REGION Network 12: IW422 - Tank Group Pressure (PT-424) - Tank Group
   RUNG wire#powerrail
      { S7_Templates := "[SrcType := Int, DestType := Real]" } Normalize(min := "20_TANKS_IP_DATA".RIO_07.FIRST_TANK.TANKS_PRESS_CNFG.RAW_MIN, value := "RIO7 Tank Pressure", max := "20_TANKS_IP_DATA".RIO_07.FIRST_TANK.TANKS_PRESS_CNFG.RAW_MAX, out => "20_TANKS_IP_DATA".RIO_07.FIRST_TANK.TANKS_PRESS_CNFG.NORM)
      { S7_Templates := "[SrcType := Real, DestType := Real]" } Scale(min := "20_TANKS_IP_DATA".RIO_07.FIRST_TANK.TANKS_PRESS_CNFG.ENG_MIN, value := "20_TANKS_IP_DATA".RIO_07.FIRST_TANK.TANKS_PRESS_CNFG.NORM, max := "20_TANKS_IP_DATA".RIO_07.FIRST_TANK.TANKS_PRESS_CNFG.ENG_MAX, out => "20_TANKS_IP_DATA".RIO_07.FIRST_TANK.TANKS_PRESS)
   END_RUNG
   // the same network as SCL:
   "20_TANKS_IP_DATA".RIO_07.FIRST_TANK.TANKS_PRESS_CNFG.NORM := NORM_X(MIN := "20_TANKS_IP_DATA".RIO_07.FIRST_TANK.TANKS_PRESS_CNFG.RAW_MIN, VALUE := "RIO7 Tank Pressure", MAX := "20_TANKS_IP_DATA".RIO_07.FIRST_TANK.TANKS_PRESS_CNFG.RAW_MAX);
   "20_TANKS_IP_DATA".RIO_07.FIRST_TANK.TANKS_PRESS := SCALE_X(MIN := "20_TANKS_IP_DATA".RIO_07.FIRST_TANK.TANKS_PRESS_CNFG.ENG_MIN, VALUE := "20_TANKS_IP_DATA".RIO_07.FIRST_TANK.TANKS_PRESS_CNFG.NORM, MAX := "20_TANKS_IP_DATA".RIO_07.FIRST_TANK.TANKS_PRESS_CNFG.ENG_MAX);
END_REGION
END_FUNCTION

FUNCTION "40_RIO_Output_Processing" : Void   // FC40, LAD
TITLE = RIO Output Processing
{ S7_Optimized_Access := 'TRUE' }
AUTHOR : JRS
VERSION : 0.1
// To call output processing blocks in logical order
BEGIN

REGION Network 1: RIO Digital Output Processing - Rack 1
   // To process code outputs prior to physical connection
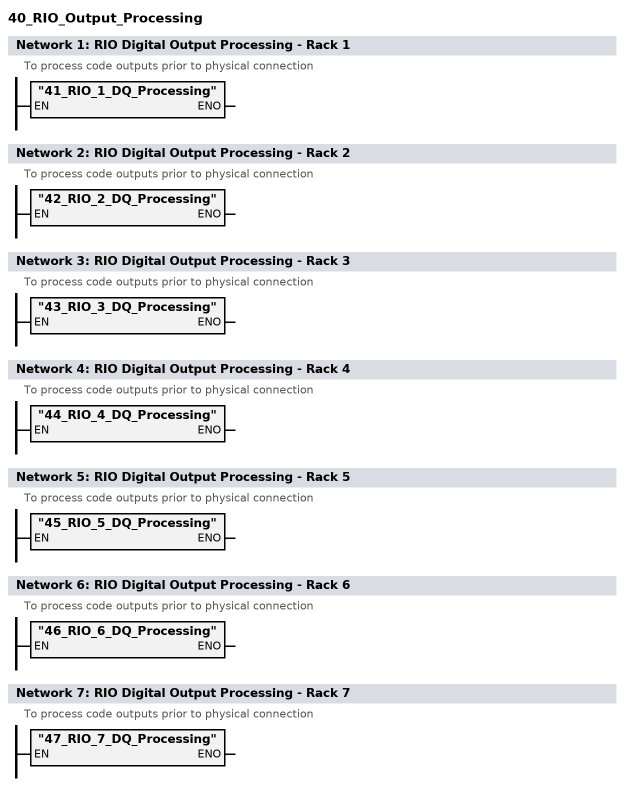
   RUNG wire#powerrail
      "41_RIO_1_DQ_Processing"()
   END_RUNG
   // the same network as SCL:
   "41_RIO_1_DQ_Processing"();
END_REGION

REGION Network 2: RIO Digital Output Processing - Rack 2
   // To process code outputs prior to physical connection
   RUNG wire#powerrail
      "42_RIO_2_DQ_Processing"()
   END_RUNG
   // the same network as SCL:
   "42_RIO_2_DQ_Processing"();
END_REGION

REGION Network 3: RIO Digital Output Processing - Rack 3
   // To process code outputs prior to physical connection
   RUNG wire#powerrail
      "43_RIO_3_DQ_Processing"()
   END_RUNG
   // the same network as SCL:
   "43_RIO_3_DQ_Processing"();
END_REGION

REGION Network 4: RIO Digital Output Processing - Rack 4
   // To process code outputs prior to physical connection
   RUNG wire#powerrail
      "44_RIO_4_DQ_Processing"()
   END_RUNG
   // the same network as SCL:
   "44_RIO_4_DQ_Processing"();
END_REGION

REGION Network 5: RIO Digital Output Processing - Rack 5
   // To process code outputs prior to physical connection
   RUNG wire#powerrail
      "45_RIO_5_DQ_Processing"()
   END_RUNG
   // the same network as SCL:
   "45_RIO_5_DQ_Processing"();
END_REGION

REGION Network 6: RIO Digital Output Processing - Rack 6
   // To process code outputs prior to physical connection
   RUNG wire#powerrail
      "46_RIO_6_DQ_Processing"()
   END_RUNG
   // the same network as SCL:
   "46_RIO_6_DQ_Processing"();
END_REGION

REGION Network 7: RIO Digital Output Processing - Rack 7
   // To process code outputs prior to physical connection
   RUNG wire#powerrail
      "47_RIO_7_DQ_Processing"()
   END_RUNG
   // the same network as SCL:
   "47_RIO_7_DQ_Processing"();
END_REGION
END_FUNCTION

FUNCTION "41_RIO_1_DQ_Processing" : Void   // FC41, LAD
TITLE = RIO Rack Digital Output Processing (Tanks APT, 1P & 1S)
{ S7_Optimized_Access := 'TRUE' }
AUTHOR : JRS
VERSION : 0.1
// To process code outputs prior to physical connection
BEGIN

REGION Network 1: Q0.0 - Tank Vent Valve Control (CV-441-A) - FPT
   // True = CLOSE, False = OPEN
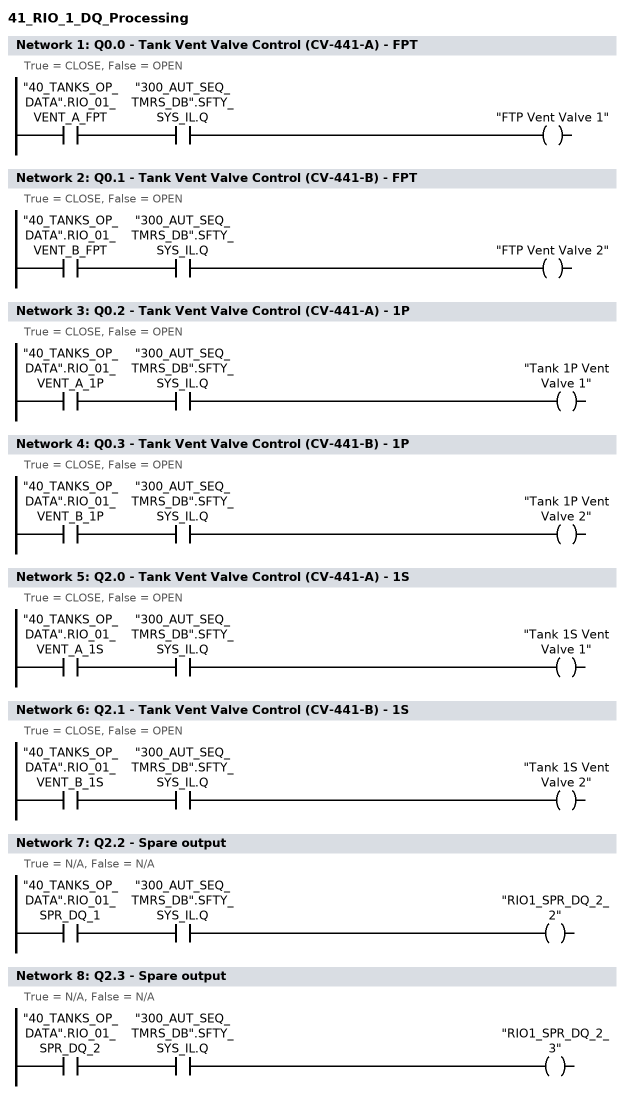
   RUNG wire#powerrail
      Contact( "40_TANKS_OP_DATA".RIO_01_VENT_A_FPT )
      Contact( "300_AUT_SEQ_TMRS_DB".SFTY_SYS_IL.Q )
      Coil( "FTP Vent Valve 1" )
   END_RUNG
   // the same network as SCL:
   "FTP Vent Valve 1" := "40_TANKS_OP_DATA".RIO_01_VENT_A_FPT AND "300_AUT_SEQ_TMRS_DB".SFTY_SYS_IL.Q;
END_REGION

REGION Network 2: Q0.1 - Tank Vent Valve Control (CV-441-B) - FPT
   // True = CLOSE, False = OPEN
   RUNG wire#powerrail
      Contact( "40_TANKS_OP_DATA".RIO_01_VENT_B_FPT )
      Contact( "300_AUT_SEQ_TMRS_DB".SFTY_SYS_IL.Q )
      Coil( "FTP Vent Valve 2" )
   END_RUNG
   // the same network as SCL:
   "FTP Vent Valve 2" := "40_TANKS_OP_DATA".RIO_01_VENT_B_FPT AND "300_AUT_SEQ_TMRS_DB".SFTY_SYS_IL.Q;
END_REGION

REGION Network 3: Q0.2 - Tank Vent Valve Control (CV-441-A) - 1P
   // True = CLOSE, False = OPEN
   RUNG wire#powerrail
      Contact( "40_TANKS_OP_DATA".RIO_01_VENT_A_1P )
      Contact( "300_AUT_SEQ_TMRS_DB".SFTY_SYS_IL.Q )
      Coil( "Tank 1P Vent Valve 1" )
   END_RUNG
   // the same network as SCL:
   "Tank 1P Vent Valve 1" := "40_TANKS_OP_DATA".RIO_01_VENT_A_1P AND "300_AUT_SEQ_TMRS_DB".SFTY_SYS_IL.Q;
END_REGION

REGION Network 4: Q0.3 - Tank Vent Valve Control (CV-441-B) - 1P
   // True = CLOSE, False = OPEN
   RUNG wire#powerrail
      Contact( "40_TANKS_OP_DATA".RIO_01_VENT_B_1P )
      Contact( "300_AUT_SEQ_TMRS_DB".SFTY_SYS_IL.Q )
      Coil( "Tank 1P Vent Valve 2" )
   END_RUNG
   // the same network as SCL:
   "Tank 1P Vent Valve 2" := "40_TANKS_OP_DATA".RIO_01_VENT_B_1P AND "300_AUT_SEQ_TMRS_DB".SFTY_SYS_IL.Q;
END_REGION

REGION Network 5: Q2.0 - Tank Vent Valve Control (CV-441-A) - 1S
   // True = CLOSE, False = OPEN
   RUNG wire#powerrail
      Contact( "40_TANKS_OP_DATA".RIO_01_VENT_A_1S )
      Contact( "300_AUT_SEQ_TMRS_DB".SFTY_SYS_IL.Q )
      Coil( "Tank 1S Vent Valve 1" )
   END_RUNG
   // the same network as SCL:
   "Tank 1S Vent Valve 1" := "40_TANKS_OP_DATA".RIO_01_VENT_A_1S AND "300_AUT_SEQ_TMRS_DB".SFTY_SYS_IL.Q;
END_REGION

REGION Network 6: Q2.1 - Tank Vent Valve Control (CV-441-B) - 1S
   // True = CLOSE, False = OPEN
   RUNG wire#powerrail
      Contact( "40_TANKS_OP_DATA".RIO_01_VENT_B_1S )
      Contact( "300_AUT_SEQ_TMRS_DB".SFTY_SYS_IL.Q )
      Coil( "Tank 1S Vent Valve 2" )
   END_RUNG
   // the same network as SCL:
   "Tank 1S Vent Valve 2" := "40_TANKS_OP_DATA".RIO_01_VENT_B_1S AND "300_AUT_SEQ_TMRS_DB".SFTY_SYS_IL.Q;
END_REGION

REGION Network 7: Q2.2 - Spare output
   // True = N/A, False = N/A
   RUNG wire#powerrail
      Contact( "40_TANKS_OP_DATA".RIO_01_SPR_DQ_1 )
      Contact( "300_AUT_SEQ_TMRS_DB".SFTY_SYS_IL.Q )
      Coil( "RIO1_SPR_DQ_2_2" )
   END_RUNG
   // the same network as SCL:
   "RIO1_SPR_DQ_2_2" := "40_TANKS_OP_DATA".RIO_01_SPR_DQ_1 AND "300_AUT_SEQ_TMRS_DB".SFTY_SYS_IL.Q;
END_REGION

REGION Network 8: Q2.3 - Spare output
   // True = N/A, False = N/A
   RUNG wire#powerrail
      Contact( "40_TANKS_OP_DATA".RIO_01_SPR_DQ_2 )
      Contact( "300_AUT_SEQ_TMRS_DB".SFTY_SYS_IL.Q )
      Coil( "RIO1_SPR_DQ_2_3" )
   END_RUNG
   // the same network as SCL:
   "RIO1_SPR_DQ_2_3" := "40_TANKS_OP_DATA".RIO_01_SPR_DQ_2 AND "300_AUT_SEQ_TMRS_DB".SFTY_SYS_IL.Q;
END_REGION
END_FUNCTION

FUNCTION "42_RIO_2_DQ_Processing" : Void   // FC42, LAD
TITLE = RIO Rack Digital Output Processing (Tanks 2P & 2S)
{ S7_Optimized_Access := 'TRUE' }
AUTHOR : JRS
VERSION : 0.1
// To process code outputs prior to physical connection
BEGIN

REGION Network 1: Q6.0 - Tank Vent Valve Control (CV-441-A) - 2P
   // True = CLOSE, False = OPEN
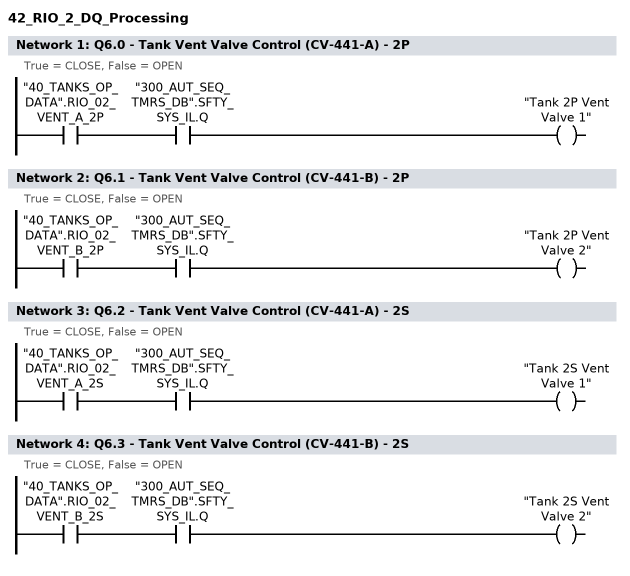
   RUNG wire#powerrail
      Contact( "40_TANKS_OP_DATA".RIO_02_VENT_A_2P )
      Contact( "300_AUT_SEQ_TMRS_DB".SFTY_SYS_IL.Q )
      Coil( "Tank 2P Vent Valve 1" )
   END_RUNG
   // the same network as SCL:
   "Tank 2P Vent Valve 1" := "40_TANKS_OP_DATA".RIO_02_VENT_A_2P AND "300_AUT_SEQ_TMRS_DB".SFTY_SYS_IL.Q;
END_REGION

REGION Network 2: Q6.1 - Tank Vent Valve Control (CV-441-B) - 2P
   // True = CLOSE, False = OPEN
   RUNG wire#powerrail
      Contact( "40_TANKS_OP_DATA".RIO_02_VENT_B_2P )
      Contact( "300_AUT_SEQ_TMRS_DB".SFTY_SYS_IL.Q )
      Coil( "Tank 2P Vent Valve 2" )
   END_RUNG
   // the same network as SCL:
   "Tank 2P Vent Valve 2" := "40_TANKS_OP_DATA".RIO_02_VENT_B_2P AND "300_AUT_SEQ_TMRS_DB".SFTY_SYS_IL.Q;
END_REGION

REGION Network 3: Q6.2 - Tank Vent Valve Control (CV-441-A) - 2S
   // True = CLOSE, False = OPEN
   RUNG wire#powerrail
      Contact( "40_TANKS_OP_DATA".RIO_02_VENT_A_2S )
      Contact( "300_AUT_SEQ_TMRS_DB".SFTY_SYS_IL.Q )
      Coil( "Tank 2S Vent Valve 1" )
   END_RUNG
   // the same network as SCL:
   "Tank 2S Vent Valve 1" := "40_TANKS_OP_DATA".RIO_02_VENT_A_2S AND "300_AUT_SEQ_TMRS_DB".SFTY_SYS_IL.Q;
END_REGION

REGION Network 4: Q6.3 - Tank Vent Valve Control (CV-441-B) - 2S
   // True = CLOSE, False = OPEN
   RUNG wire#powerrail
      Contact( "40_TANKS_OP_DATA".RIO_02_VENT_B_2S )
      Contact( "300_AUT_SEQ_TMRS_DB".SFTY_SYS_IL.Q )
      Coil( "Tank 2S Vent Valve 2" )
   END_RUNG
   // the same network as SCL:
   "Tank 2S Vent Valve 2" := "40_TANKS_OP_DATA".RIO_02_VENT_B_2S AND "300_AUT_SEQ_TMRS_DB".SFTY_SYS_IL.Q;
END_REGION
END_FUNCTION

FUNCTION "43_RIO_3_DQ_Processing" : Void   // FC43, LAD
TITLE = RIO Rack Digital Output Processing (Tanks 3P & 3S)
{ S7_Optimized_Access := 'TRUE' }
AUTHOR : JRS
VERSION : 0.1
// To process code outputs prior to physical connection
BEGIN

REGION Network 1: Q10.0 - Tank Vent Valve Control (CV-441-A) - 3P
   // True = CLOSE, False = OPEN
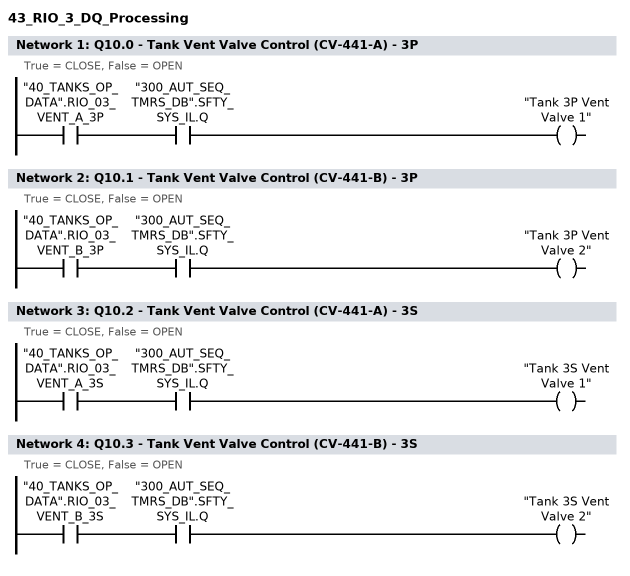
   RUNG wire#powerrail
      Contact( "40_TANKS_OP_DATA".RIO_03_VENT_A_3P )
      Contact( "300_AUT_SEQ_TMRS_DB".SFTY_SYS_IL.Q )
      Coil( "Tank 3P Vent Valve 1" )
   END_RUNG
   // the same network as SCL:
   "Tank 3P Vent Valve 1" := "40_TANKS_OP_DATA".RIO_03_VENT_A_3P AND "300_AUT_SEQ_TMRS_DB".SFTY_SYS_IL.Q;
END_REGION

REGION Network 2: Q10.1 - Tank Vent Valve Control (CV-441-B) - 3P
   // True = CLOSE, False = OPEN
   RUNG wire#powerrail
      Contact( "40_TANKS_OP_DATA".RIO_03_VENT_B_3P )
      Contact( "300_AUT_SEQ_TMRS_DB".SFTY_SYS_IL.Q )
      Coil( "Tank 3P Vent Valve 2" )
   END_RUNG
   // the same network as SCL:
   "Tank 3P Vent Valve 2" := "40_TANKS_OP_DATA".RIO_03_VENT_B_3P AND "300_AUT_SEQ_TMRS_DB".SFTY_SYS_IL.Q;
END_REGION

REGION Network 3: Q10.2 - Tank Vent Valve Control (CV-441-A) - 3S
   // True = CLOSE, False = OPEN
   RUNG wire#powerrail
      Contact( "40_TANKS_OP_DATA".RIO_03_VENT_A_3S )
      Contact( "300_AUT_SEQ_TMRS_DB".SFTY_SYS_IL.Q )
      Coil( "Tank 3S Vent Valve 1" )
   END_RUNG
   // the same network as SCL:
   "Tank 3S Vent Valve 1" := "40_TANKS_OP_DATA".RIO_03_VENT_A_3S AND "300_AUT_SEQ_TMRS_DB".SFTY_SYS_IL.Q;
END_REGION

REGION Network 4: Q10.3 - Tank Vent Valve Control (CV-441-B) - 3S
   // True = CLOSE, False = OPEN
   RUNG wire#powerrail
      Contact( "40_TANKS_OP_DATA".RIO_03_VENT_B_3S )
      Contact( "300_AUT_SEQ_TMRS_DB".SFTY_SYS_IL.Q )
      Coil( "Tank 3S Vent Valve 2" )
   END_RUNG
   // the same network as SCL:
   "Tank 3S Vent Valve 2" := "40_TANKS_OP_DATA".RIO_03_VENT_B_3S AND "300_AUT_SEQ_TMRS_DB".SFTY_SYS_IL.Q;
END_REGION
END_FUNCTION

FUNCTION "44_RIO_4_DQ_Processing" : Void   // FC44, LAD
TITLE = RIO Rack Digital Output Processing (Tanks 4P & 4S)
{ S7_Optimized_Access := 'TRUE' }
AUTHOR : JRS
VERSION : 0.1
// To process code outputs prior to physical connection
BEGIN

REGION Network 1: Q14.0 - Tank Vent Valve Control (CV-441-A) - 4P
   // True = CLOSE, False = OPEN
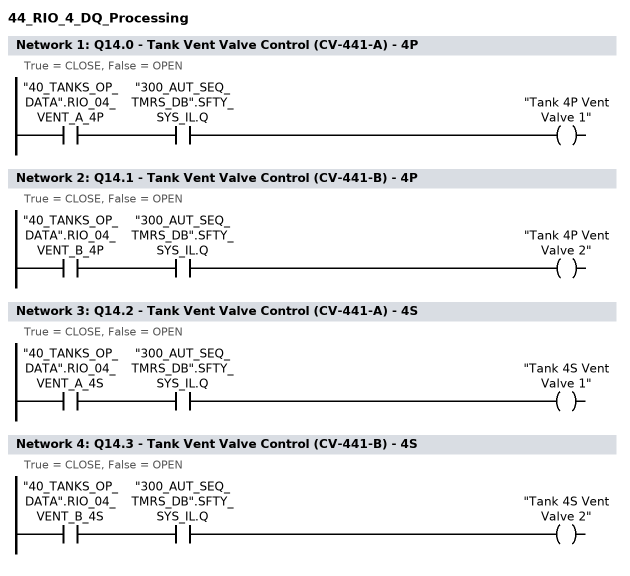
   RUNG wire#powerrail
      Contact( "40_TANKS_OP_DATA".RIO_04_VENT_A_4P )
      Contact( "300_AUT_SEQ_TMRS_DB".SFTY_SYS_IL.Q )
      Coil( "Tank 4P Vent Valve 1" )
   END_RUNG
   // the same network as SCL:
   "Tank 4P Vent Valve 1" := "40_TANKS_OP_DATA".RIO_04_VENT_A_4P AND "300_AUT_SEQ_TMRS_DB".SFTY_SYS_IL.Q;
END_REGION

REGION Network 2: Q14.1 - Tank Vent Valve Control (CV-441-B) - 4P
   // True = CLOSE, False = OPEN
   RUNG wire#powerrail
      Contact( "40_TANKS_OP_DATA".RIO_04_VENT_B_4P )
      Contact( "300_AUT_SEQ_TMRS_DB".SFTY_SYS_IL.Q )
      Coil( "Tank 4P Vent Valve 2" )
   END_RUNG
   // the same network as SCL:
   "Tank 4P Vent Valve 2" := "40_TANKS_OP_DATA".RIO_04_VENT_B_4P AND "300_AUT_SEQ_TMRS_DB".SFTY_SYS_IL.Q;
END_REGION

REGION Network 3: Q14.2 - Tank Vent Valve Control (CV-441-A) - 4S
   // True = CLOSE, False = OPEN
   RUNG wire#powerrail
      Contact( "40_TANKS_OP_DATA".RIO_04_VENT_A_4S )
      Contact( "300_AUT_SEQ_TMRS_DB".SFTY_SYS_IL.Q )
      Coil( "Tank 4S Vent Valve 1" )
   END_RUNG
   // the same network as SCL:
   "Tank 4S Vent Valve 1" := "40_TANKS_OP_DATA".RIO_04_VENT_A_4S AND "300_AUT_SEQ_TMRS_DB".SFTY_SYS_IL.Q;
END_REGION

REGION Network 4: Q14.3 - Tank Vent Valve Control (CV-441-B) - 4S
   // True = CLOSE, False = OPEN
   RUNG wire#powerrail
      Contact( "40_TANKS_OP_DATA".RIO_04_VENT_B_4S )
      Contact( "300_AUT_SEQ_TMRS_DB".SFTY_SYS_IL.Q )
      Coil( "Tank 4S Vent Valve 2" )
   END_RUNG
   // the same network as SCL:
   "Tank 4S Vent Valve 2" := "40_TANKS_OP_DATA".RIO_04_VENT_B_4S AND "300_AUT_SEQ_TMRS_DB".SFTY_SYS_IL.Q;
END_REGION
END_FUNCTION

FUNCTION "45_RIO_5_DQ_Processing" : Void   // FC45, LAD
TITLE = RIO Rack Digital Output Processing (Tanks 5P & 5S)
{ S7_Optimized_Access := 'TRUE' }
AUTHOR : JRS
VERSION : 0.1
// To process code outputs prior to physical connection
BEGIN

REGION Network 1: Q18.0 - Tank Vent Valve Control (CV-441-A) - 5P
   // True = CLOSE, False = OPEN
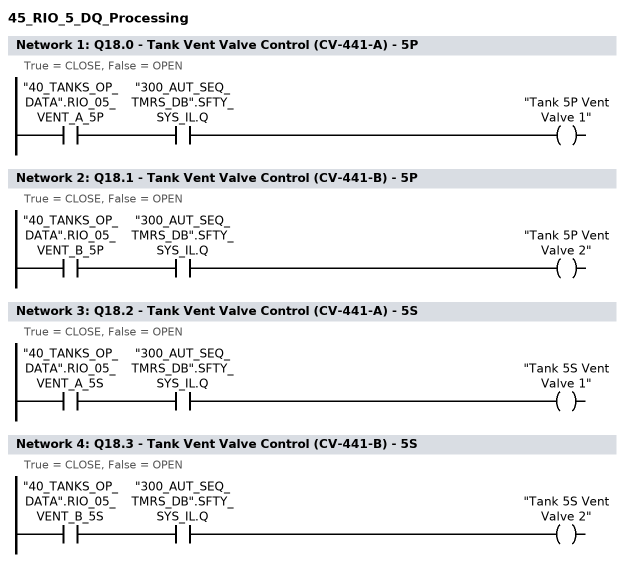
   RUNG wire#powerrail
      Contact( "40_TANKS_OP_DATA".RIO_05_VENT_A_5P )
      Contact( "300_AUT_SEQ_TMRS_DB".SFTY_SYS_IL.Q )
      Coil( "Tank 5P Vent Valve 1" )
   END_RUNG
   // the same network as SCL:
   "Tank 5P Vent Valve 1" := "40_TANKS_OP_DATA".RIO_05_VENT_A_5P AND "300_AUT_SEQ_TMRS_DB".SFTY_SYS_IL.Q;
END_REGION

REGION Network 2: Q18.1 - Tank Vent Valve Control (CV-441-B) - 5P
   // True = CLOSE, False = OPEN
   RUNG wire#powerrail
      Contact( "40_TANKS_OP_DATA".RIO_05_VENT_B_5P )
      Contact( "300_AUT_SEQ_TMRS_DB".SFTY_SYS_IL.Q )
      Coil( "Tank 5P Vent Valve 2" )
   END_RUNG
   // the same network as SCL:
   "Tank 5P Vent Valve 2" := "40_TANKS_OP_DATA".RIO_05_VENT_B_5P AND "300_AUT_SEQ_TMRS_DB".SFTY_SYS_IL.Q;
END_REGION

REGION Network 3: Q18.2 - Tank Vent Valve Control (CV-441-A) - 5S
   // True = CLOSE, False = OPEN
   RUNG wire#powerrail
      Contact( "40_TANKS_OP_DATA".RIO_05_VENT_A_5S )
      Contact( "300_AUT_SEQ_TMRS_DB".SFTY_SYS_IL.Q )
      Coil( "Tank 5S Vent Valve 1" )
   END_RUNG
   // the same network as SCL:
   "Tank 5S Vent Valve 1" := "40_TANKS_OP_DATA".RIO_05_VENT_A_5S AND "300_AUT_SEQ_TMRS_DB".SFTY_SYS_IL.Q;
END_REGION

REGION Network 4: Q18.3 - Tank Vent Valve Control (CV-441-B) - 5S
   // True = CLOSE, False = OPEN
   RUNG wire#powerrail
      Contact( "40_TANKS_OP_DATA".RIO_05_VENT_B_5S )
      Contact( "300_AUT_SEQ_TMRS_DB".SFTY_SYS_IL.Q )
      Coil( "Tank 5S Vent Valve 2" )
   END_RUNG
   // the same network as SCL:
   "Tank 5S Vent Valve 2" := "40_TANKS_OP_DATA".RIO_05_VENT_B_5S AND "300_AUT_SEQ_TMRS_DB".SFTY_SYS_IL.Q;
END_REGION
END_FUNCTION

FUNCTION "46_RIO_6_DQ_Processing" : Void   // FC46, LAD
TITLE = RIO Rack Digital Output Processing (Tanks 6P & 6S)
{ S7_Optimized_Access := 'TRUE' }
AUTHOR : JRS
VERSION : 0.1
// To process code outputs prior to physical connection
BEGIN

REGION Network 1: Q20.0 - Tank Vent Valve Control (CV-441-A) - 6P
   // True = CLOSE, False = OPEN
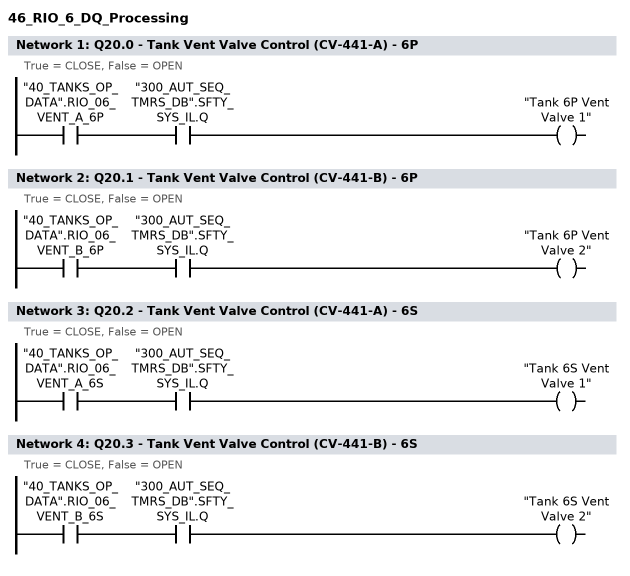
   RUNG wire#powerrail
      Contact( "40_TANKS_OP_DATA".RIO_06_VENT_A_6P )
      Contact( "300_AUT_SEQ_TMRS_DB".SFTY_SYS_IL.Q )
      Coil( "Tank 6P Vent Valve 1" )
   END_RUNG
   // the same network as SCL:
   "Tank 6P Vent Valve 1" := "40_TANKS_OP_DATA".RIO_06_VENT_A_6P AND "300_AUT_SEQ_TMRS_DB".SFTY_SYS_IL.Q;
END_REGION

REGION Network 2: Q20.1 - Tank Vent Valve Control (CV-441-B) - 6P
   // True = CLOSE, False = OPEN
   RUNG wire#powerrail
      Contact( "40_TANKS_OP_DATA".RIO_06_VENT_B_6P )
      Contact( "300_AUT_SEQ_TMRS_DB".SFTY_SYS_IL.Q )
      Coil( "Tank 6P Vent Valve 2" )
   END_RUNG
   // the same network as SCL:
   "Tank 6P Vent Valve 2" := "40_TANKS_OP_DATA".RIO_06_VENT_B_6P AND "300_AUT_SEQ_TMRS_DB".SFTY_SYS_IL.Q;
END_REGION

REGION Network 3: Q20.2 - Tank Vent Valve Control (CV-441-A) - 6S
   // True = CLOSE, False = OPEN
   RUNG wire#powerrail
      Contact( "40_TANKS_OP_DATA".RIO_06_VENT_A_6S )
      Contact( "300_AUT_SEQ_TMRS_DB".SFTY_SYS_IL.Q )
      Coil( "Tank 6S Vent Valve 1" )
   END_RUNG
   // the same network as SCL:
   "Tank 6S Vent Valve 1" := "40_TANKS_OP_DATA".RIO_06_VENT_A_6S AND "300_AUT_SEQ_TMRS_DB".SFTY_SYS_IL.Q;
END_REGION

REGION Network 4: Q20.3 - Tank Vent Valve Control (CV-441-B) - 6S
   // True = CLOSE, False = OPEN
   RUNG wire#powerrail
      Contact( "40_TANKS_OP_DATA".RIO_06_VENT_B_6S )
      Contact( "300_AUT_SEQ_TMRS_DB".SFTY_SYS_IL.Q )
      Coil( "Tank 6S Vent Valve 2" )
   END_RUNG
   // the same network as SCL:
   "Tank 6S Vent Valve 2" := "40_TANKS_OP_DATA".RIO_06_VENT_B_6S AND "300_AUT_SEQ_TMRS_DB".SFTY_SYS_IL.Q;
END_REGION
END_FUNCTION

FUNCTION "47_RIO_7_DQ_Processing" : Void   // FC47, LAD
TITLE = RIO Rack Digital Output Processing (Tank APT)
{ S7_Optimized_Access := 'TRUE' }
AUTHOR : JRS
VERSION : 0.1
// To process code outputs prior to physical connection
BEGIN

REGION Network 1: Q26.0 - Tank Vent Valve Control (CV-441-A) - APT
   // True = CLOSE, False = OPEN
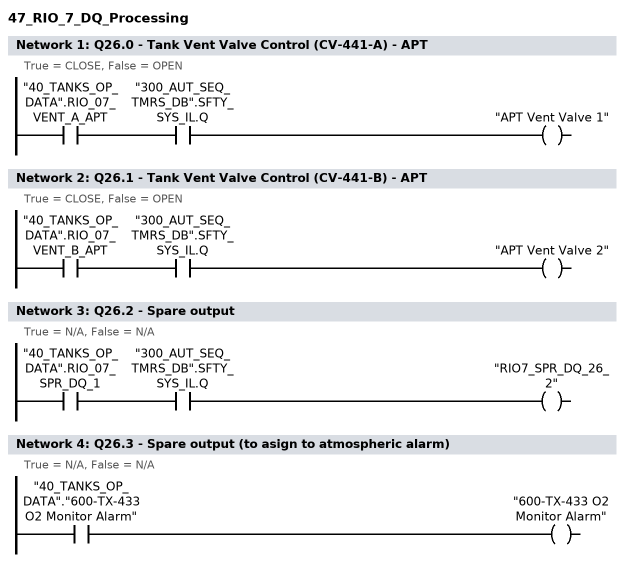
   RUNG wire#powerrail
      Contact( "40_TANKS_OP_DATA".RIO_07_VENT_A_APT )
      Contact( "300_AUT_SEQ_TMRS_DB".SFTY_SYS_IL.Q )
      Coil( "APT Vent Valve 1" )
   END_RUNG
   // the same network as SCL:
   "APT Vent Valve 1" := "40_TANKS_OP_DATA".RIO_07_VENT_A_APT AND "300_AUT_SEQ_TMRS_DB".SFTY_SYS_IL.Q;
END_REGION

REGION Network 2: Q26.1 - Tank Vent Valve Control (CV-441-B) - APT
   // True = CLOSE, False = OPEN
   RUNG wire#powerrail
      Contact( "40_TANKS_OP_DATA".RIO_07_VENT_B_APT )
      Contact( "300_AUT_SEQ_TMRS_DB".SFTY_SYS_IL.Q )
      Coil( "APT Vent Valve 2" )
   END_RUNG
   // the same network as SCL:
   "APT Vent Valve 2" := "40_TANKS_OP_DATA".RIO_07_VENT_B_APT AND "300_AUT_SEQ_TMRS_DB".SFTY_SYS_IL.Q;
END_REGION

REGION Network 3: Q26.2 - Spare output
   // True = N/A, False = N/A
   RUNG wire#powerrail
      Contact( "40_TANKS_OP_DATA".RIO_07_SPR_DQ_1 )
      Contact( "300_AUT_SEQ_TMRS_DB".SFTY_SYS_IL.Q )
      Coil( "RIO7_SPR_DQ_26_2" )
   END_RUNG
   // the same network as SCL:
   "RIO7_SPR_DQ_26_2" := "40_TANKS_OP_DATA".RIO_07_SPR_DQ_1 AND "300_AUT_SEQ_TMRS_DB".SFTY_SYS_IL.Q;
END_REGION

REGION Network 4: Q26.3 - Spare output (to asign to atmospheric alarm)
   // True = N/A, False = N/A
   RUNG wire#powerrail
      Contact( "40_TANKS_OP_DATA"."600-TX-433  O2 Monitor Alarm" )
      Coil( "600-TX-433 O2 Monitor Alarm" )
   END_RUNG
   // the same network as SCL:
   "600-TX-433 O2 Monitor Alarm" := "40_TANKS_OP_DATA"."600-TX-433  O2 Monitor Alarm";
END_REGION
END_FUNCTION

// folder: 2000 - 2999 BTCS System/2010 - 2019 IO & Processing

FUNCTION_BLOCK "2019_Tank_Auto_Cmds"   // FB2019, LAD
{ S7_Optimized_Access := 'TRUE' }
VERSION : 0.1
   VAR_INPUT
      Run : Bool;
   END_VAR
BEGIN

REGION Network 2: Q136.2 - Block Valve 1 Control (CV407) +++Control By BWTS+++ N.C.
   // True = OPEN, False = CLOSE
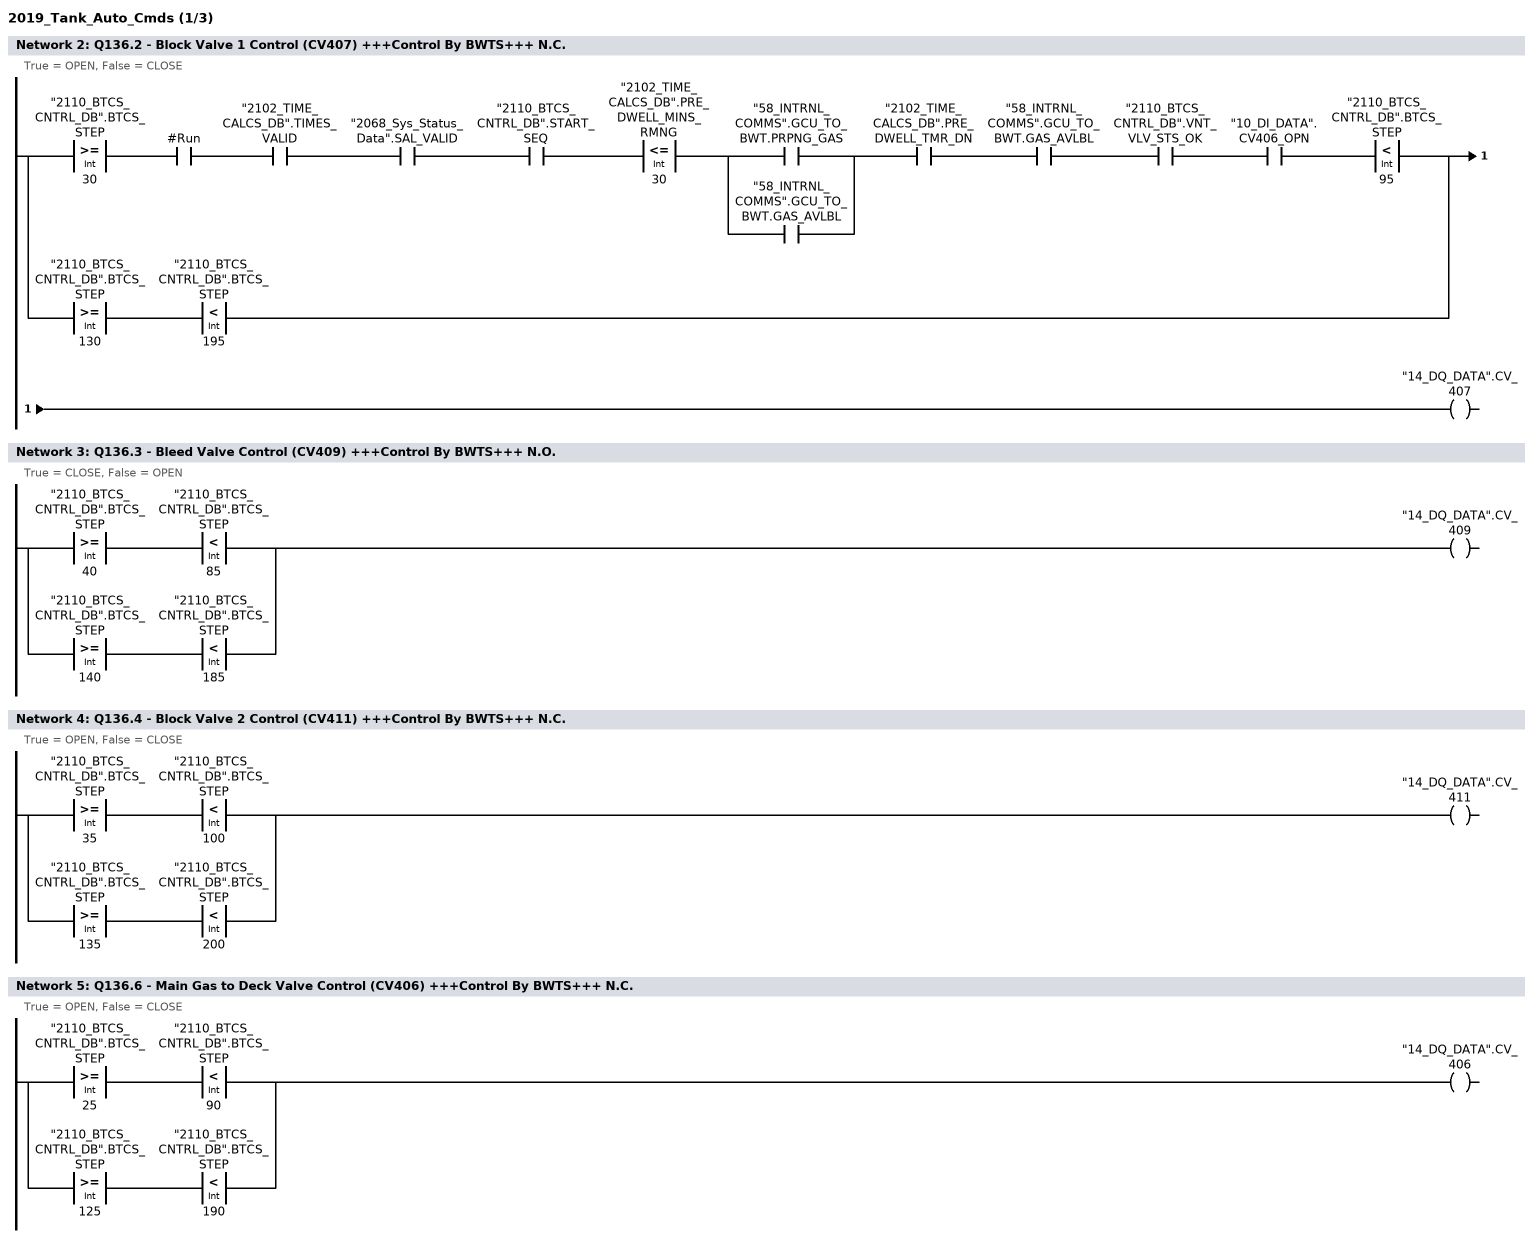
   RUNG wire#powerrail
      { S7_Templates := "SrcType := Int" } GE_Contact(in1 := "2110_BTCS_CNTRL_DB".BTCS_STEP, in2 := 30)
      Contact( #Run )
      Contact( "2102_TIME_CALCS_DB".TIMES_VALID )
      Contact( "2068_Sys_Status_Data".SAL_VALID )
      Contact( "2110_BTCS_CNTRL_DB".START_SEQ )
      { S7_Templates := "SrcType := Int" } LE_Contact(in1 := "2102_TIME_CALCS_DB".PRE_DWELL_MINS_RMNG, in2 := 30)
      wire#w1
      Contact( "58_INTRNL_COMMS".GCU_TO_BWT.PRPNG_GAS )
      wire#w2
      Contact( "2102_TIME_CALCS_DB".PRE_DWELL_TMR_DN )
      Contact( "58_INTRNL_COMMS".GCU_TO_BWT.GAS_AVLBL )
      Contact( "2110_BTCS_CNTRL_DB".VNT_VLV_STS_OK )
      Contact( "10_DI_DATA".CV406_OPN )
      { S7_Templates := "SrcType := Int" } LT_Contact(in1 := "2110_BTCS_CNTRL_DB".BTCS_STEP, in2 := 95)
      wire#w3
      Coil( "14_DQ_DATA".CV_407 )
   END_RUNG
   RUNG wire#w1
      Contact( "58_INTRNL_COMMS".GCU_TO_BWT.GAS_AVLBL )
   END_RUNG wire#w2
   RUNG wire#powerrail
      { S7_Templates := "SrcType := Int" } GE_Contact(in1 := "2110_BTCS_CNTRL_DB".BTCS_STEP, in2 := 130)
      { S7_Templates := "SrcType := Int" } LT_Contact(in1 := "2110_BTCS_CNTRL_DB".BTCS_STEP, in2 := 195)
   END_RUNG wire#w3
   // the same network as SCL:
   "14_DQ_DATA".CV_407 := (("2110_BTCS_CNTRL_DB".BTCS_STEP >= 30) AND #Run AND "2102_TIME_CALCS_DB".TIMES_VALID AND "2068_Sys_Status_Data".SAL_VALID AND "2110_BTCS_CNTRL_DB".START_SEQ AND ("2102_TIME_CALCS_DB".PRE_DWELL_MINS_RMNG <= 30) AND ("58_INTRNL_COMMS".GCU_TO_BWT.PRPNG_GAS OR "58_INTRNL_COMMS".GCU_TO_BWT.GAS_AVLBL) AND "2102_TIME_CALCS_DB".PRE_DWELL_TMR_DN AND "58_INTRNL_COMMS".GCU_TO_BWT.GAS_AVLBL AND "2110_BTCS_CNTRL_DB".VNT_VLV_STS_OK AND "10_DI_DATA".CV406_OPN AND ("2110_BTCS_CNTRL_DB".BTCS_STEP < 95)) OR (("2110_BTCS_CNTRL_DB".BTCS_STEP >= 130) AND ("2110_BTCS_CNTRL_DB".BTCS_STEP < 195));
END_REGION

REGION Network 3: Q136.3 - Bleed Valve Control (CV409) +++Control By BWTS+++ N.O.
   // True = CLOSE, False = OPEN
   RUNG wire#powerrail
      { S7_Templates := "SrcType := Int" } GE_Contact(in1 := "2110_BTCS_CNTRL_DB".BTCS_STEP, in2 := 40)
      { S7_Templates := "SrcType := Int" } LT_Contact(in1 := "2110_BTCS_CNTRL_DB".BTCS_STEP, in2 := 85)
      wire#w1
      Coil( "14_DQ_DATA".CV_409 )
   END_RUNG
   RUNG wire#powerrail
      { S7_Templates := "SrcType := Int" } GE_Contact(in1 := "2110_BTCS_CNTRL_DB".BTCS_STEP, in2 := 140)
      { S7_Templates := "SrcType := Int" } LT_Contact(in1 := "2110_BTCS_CNTRL_DB".BTCS_STEP, in2 := 185)
   END_RUNG wire#w1
   // the same network as SCL:
   "14_DQ_DATA".CV_409 := (("2110_BTCS_CNTRL_DB".BTCS_STEP >= 40) AND ("2110_BTCS_CNTRL_DB".BTCS_STEP < 85)) OR (("2110_BTCS_CNTRL_DB".BTCS_STEP >= 140) AND ("2110_BTCS_CNTRL_DB".BTCS_STEP < 185));
END_REGION

REGION Network 4: Q136.4 - Block Valve 2 Control (CV411) +++Control By BWTS+++ N.C.
   // True = OPEN, False = CLOSE
   RUNG wire#powerrail
      { S7_Templates := "SrcType := Int" } GE_Contact(in1 := "2110_BTCS_CNTRL_DB".BTCS_STEP, in2 := 35)
      { S7_Templates := "SrcType := Int" } LT_Contact(in1 := "2110_BTCS_CNTRL_DB".BTCS_STEP, in2 := 100)
      wire#w1
      Coil( "14_DQ_DATA".CV_411 )
   END_RUNG
   RUNG wire#powerrail
      { S7_Templates := "SrcType := Int" } GE_Contact(in1 := "2110_BTCS_CNTRL_DB".BTCS_STEP, in2 := 135)
      { S7_Templates := "SrcType := Int" } LT_Contact(in1 := "2110_BTCS_CNTRL_DB".BTCS_STEP, in2 := 200)
   END_RUNG wire#w1
   // the same network as SCL:
   "14_DQ_DATA".CV_411 := (("2110_BTCS_CNTRL_DB".BTCS_STEP >= 35) AND ("2110_BTCS_CNTRL_DB".BTCS_STEP < 100)) OR (("2110_BTCS_CNTRL_DB".BTCS_STEP >= 135) AND ("2110_BTCS_CNTRL_DB".BTCS_STEP < 200));
END_REGION

REGION Network 5: Q136.6 - Main Gas to Deck Valve Control (CV406) +++Control By BWTS+++ N.C.
   // True = OPEN, False = CLOSE
   RUNG wire#powerrail
      { S7_Templates := "SrcType := Int" } GE_Contact(in1 := "2110_BTCS_CNTRL_DB".BTCS_STEP, in2 := 25)
      { S7_Templates := "SrcType := Int" } LT_Contact(in1 := "2110_BTCS_CNTRL_DB".BTCS_STEP, in2 := 90)
      wire#w1
      Coil( "14_DQ_DATA".CV_406 )
   END_RUNG
   RUNG wire#powerrail
      { S7_Templates := "SrcType := Int" } GE_Contact(in1 := "2110_BTCS_CNTRL_DB".BTCS_STEP, in2 := 125)
      { S7_Templates := "SrcType := Int" } LT_Contact(in1 := "2110_BTCS_CNTRL_DB".BTCS_STEP, in2 := 190)
   END_RUNG wire#w1
   // the same network as SCL:
   "14_DQ_DATA".CV_406 := (("2110_BTCS_CNTRL_DB".BTCS_STEP >= 25) AND ("2110_BTCS_CNTRL_DB".BTCS_STEP < 90)) OR (("2110_BTCS_CNTRL_DB".BTCS_STEP >= 125) AND ("2110_BTCS_CNTRL_DB".BTCS_STEP < 190));
END_REGION

REGION Network 6: Q138.3 - Pilot For GTT 2 Port Valve (CV422-2P) +++Control By BWTS+++ N.C.
   // True = OPEN, False = CLOSE